(* Logix 5000 project; controller PLC_MCC1300_75F1 vendor 1 type 14 code 166 rev 32.11; software revision 32.04; part 16 of 83 *)
(* tags used below, declared in another part *)
   M302SpeedUp : MAC_SpeedUp;
   TMP_d : DINT;
   TMP_xPositioning : BOOL;
   TMP_xReverse : BOOL;
   TMP_xRun : BOOL;
   xAlwaysOFF : BOOL;
   Z300_Conveyor : UDT_StandConv[29];
   Z300_Conveyor_Conf : UDT_Conveyor_Config[29];
   Z300_Conveyor_HMW : MAC_Conveyor_ZC_HMW[29];
   Z300_Conveyor_IN_MOTION : MAC_Conveyor_ZC_IN_MOTION[29];
   Z301_HMR : MAC_Zone_ML_HMR;
(* CommandLogic, continued *)

ROUTINE M307AM2_Conveyor_Output   (* ladder *)
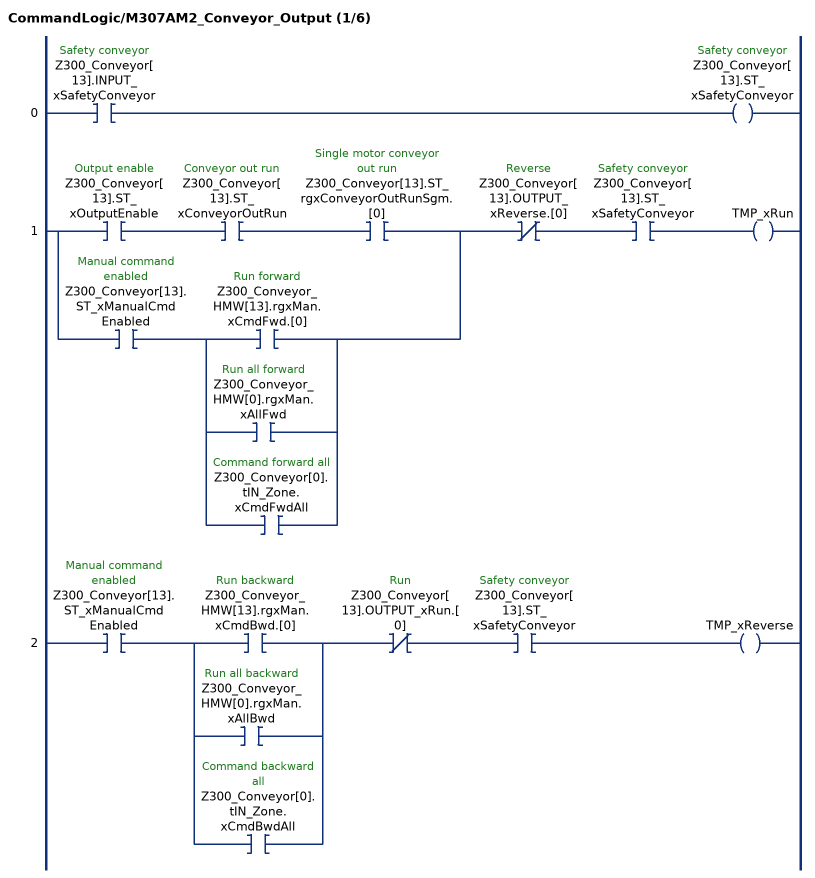
   0: XIC(Z300_Conveyor[13].INPUT_xSafetyConveyor)OTE(Z300_Conveyor[13].ST_xSafetyConveyor);
   1: [XIC(Z300_Conveyor[13].ST_xOutputEnable) XIC(Z300_Conveyor[13].ST_xConveyorOutRun) XIC(Z300_Conveyor[13].ST_rgxConveyorOutRunSgm.[0]) ,XIC(Z300_Conveyor[13].ST_xManualCmdEnabled) [XIC(Z300_Conveyor_HMW[13].rgxMan.xCmdFwd.[0]) ,XIC(Z300_Conveyor_HMW[0].rgxMan.xAllFwd) ,XIC(Z300_Conveyor[0].tIN_Zone.xCmdFwdAll) ] ]XIO(Z300_Conveyor[13].OUTPUT_xReverse.[0])XIC(Z300_Conveyor[13].ST_xSafetyConveyor)OTE(TMP_xRun);
   2: XIC(Z300_Conveyor[13].ST_xManualCmdEnabled)[XIC(Z300_Conveyor_HMW[13].rgxMan.xCmdBwd.[0]) ,XIC(Z300_Conveyor_HMW[0].rgxMan.xAllBwd) ,XIC(Z300_Conveyor[0].tIN_Zone.xCmdBwdAll) ]XIO(Z300_Conveyor[13].OUTPUT_xRun.[0])XIC(Z300_Conveyor[13].ST_xSafetyConveyor)OTE(TMP_xReverse);
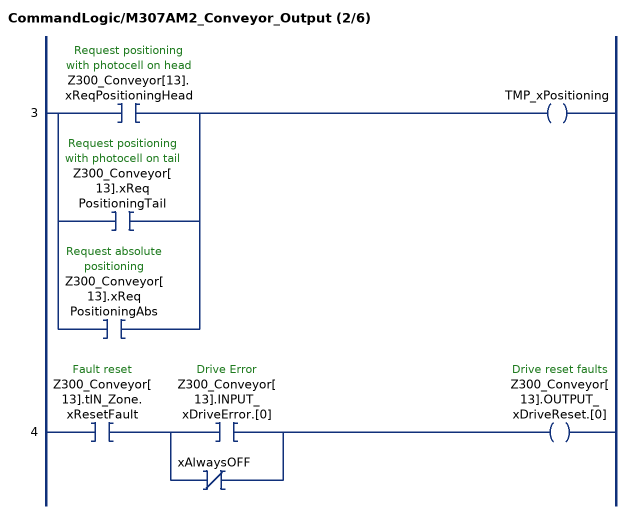
   3: [XIC(Z300_Conveyor[13].xReqPositioningHead) ,XIC(Z300_Conveyor[13].xReqPositioningTail) ,XIC(Z300_Conveyor[13].xReqPositioningAbs) ]OTE(TMP_xPositioning);
   4: XIC(Z300_Conveyor[13].tIN_Zone.xResetFault)[XIC(Z300_Conveyor[13].INPUT_xDriveError.[0]) ,XIO(xAlwaysOFF) ]OTE(Z300_Conveyor[13].OUTPUT_xDriveReset.[0]);
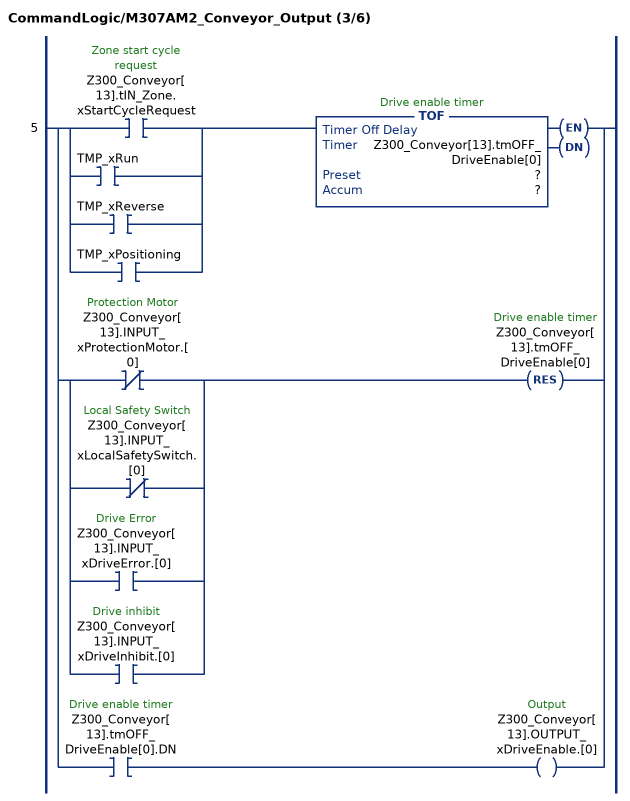
   5: [[XIC(Z300_Conveyor[13].tIN_Zone.xStartCycleRequest) ,XIC(TMP_xRun) ,XIC(TMP_xReverse) ,XIC(TMP_xPositioning) ] TOF(Z300_Conveyor[13].tmOFF_DriveEnable[0],?,?) ,[XIO(Z300_Conveyor[13].INPUT_xProtectionMotor.[0]) ,XIO(Z300_Conveyor[13].INPUT_xLocalSafetySwitch.[0]) ,XIC(Z300_Conveyor[13].INPUT_xDriveError.[0]) ,XIC(Z300_Conveyor[13].INPUT_xDriveInhibit.[0]) ] RES(Z300_Conveyor[13].tmOFF_DriveEnable[0]) ,XIC(Z300_Conveyor[13].tmOFF_DriveEnable[0].DN) OTE(Z300_Conveyor[13].OUTPUT_xDriveEnable.[0]) ];
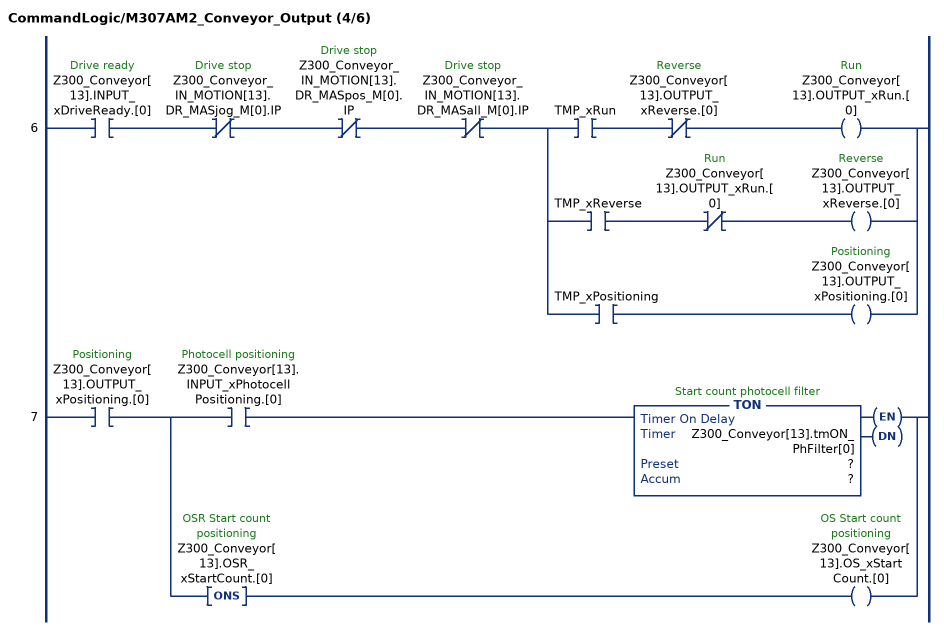
   6: XIC(Z300_Conveyor[13].INPUT_xDriveReady.[0])XIO(Z300_Conveyor_IN_MOTION[13].DR_MASjog_M[0].IP)XIO(Z300_Conveyor_IN_MOTION[13].DR_MASpos_M[0].IP)XIO(Z300_Conveyor_IN_MOTION[13].DR_MASall_M[0].IP)[XIC(TMP_xRun) XIO(Z300_Conveyor[13].OUTPUT_xReverse.[0]) OTE(Z300_Conveyor[13].OUTPUT_xRun.[0]) ,XIC(TMP_xReverse) XIO(Z300_Conveyor[13].OUTPUT_xRun.[0]) OTE(Z300_Conveyor[13].OUTPUT_xReverse.[0]) ,XIC(TMP_xPositioning) OTE(Z300_Conveyor[13].OUTPUT_xPositioning.[0]) ];
   7: XIC(Z300_Conveyor[13].OUTPUT_xPositioning.[0])[XIC(Z300_Conveyor[13].INPUT_xPhotocellPositioning.[0]) TON(Z300_Conveyor[13].tmON_PhFilter[0],?,?) ,ONS(Z300_Conveyor[13].OSR_xStartCount.[0]) OTE(Z300_Conveyor[13].OS_xStartCount.[0]) ];
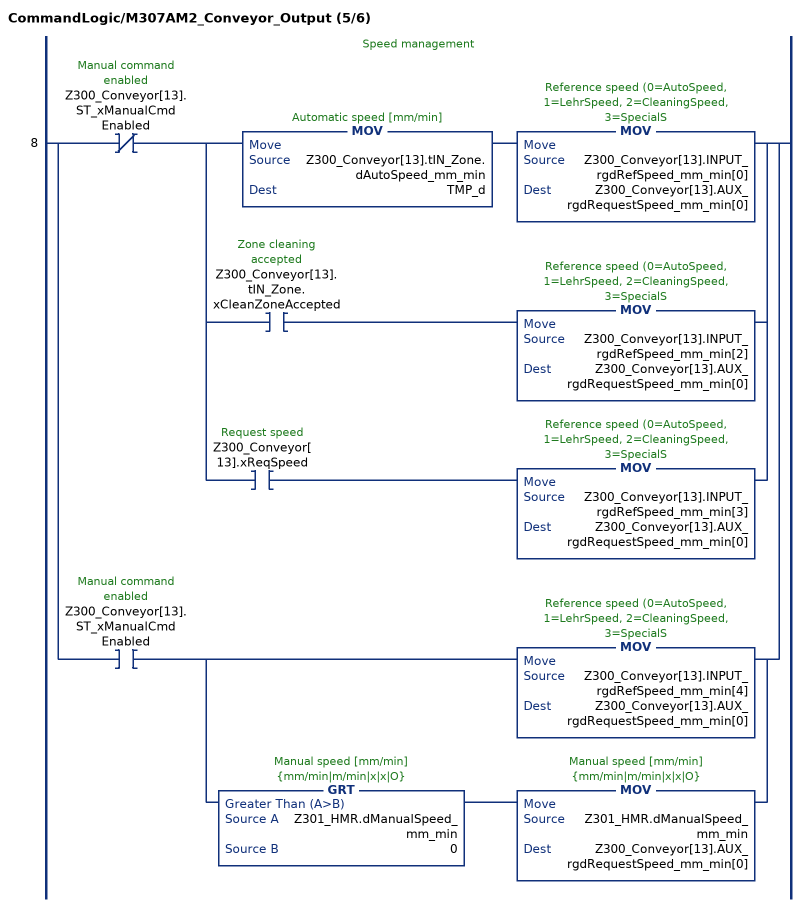
   // Speed management
   8: [XIO(Z300_Conveyor[13].ST_xManualCmdEnabled) [MOV(Z300_Conveyor[13].tIN_Zone.dAutoSpeed_mm_min,TMP_d) MOV(Z300_Conveyor[13].INPUT_rgdRefSpeed_mm_min[0],Z300_Conveyor[13].AUX_rgdRequestSpeed_mm_min[0]) ,XIC(Z300_Conveyor[13].tIN_Zone.xCleanZoneAccepted) MOV(Z300_Conveyor[13].INPUT_rgdRefSpeed_mm_min[2],Z300_Conveyor[13].AUX_rgdRequestSpeed_mm_min[0]) ,XIC(Z300_Conveyor[13].xReqSpeed) MOV(Z300_Conveyor[13].INPUT_rgdRefSpeed_mm_min[3],Z300_Conveyor[13].AUX_rgdRequestSpeed_mm_min[0]) ] ,XIC(Z300_Conveyor[13].ST_xManualCmdEnabled) [MOV(Z300_Conveyor[13].INPUT_rgdRefSpeed_mm_min[4],Z300_Conveyor[13].AUX_rgdRequestSpeed_mm_min[0]) ,GRT(Z301_HMR.dManualSpeed_mm_min,0) MOV(Z301_HMR.dManualSpeed_mm_min,Z300_Conveyor[13].AUX_rgdRequestSpeed_mm_min[0]) ] ];
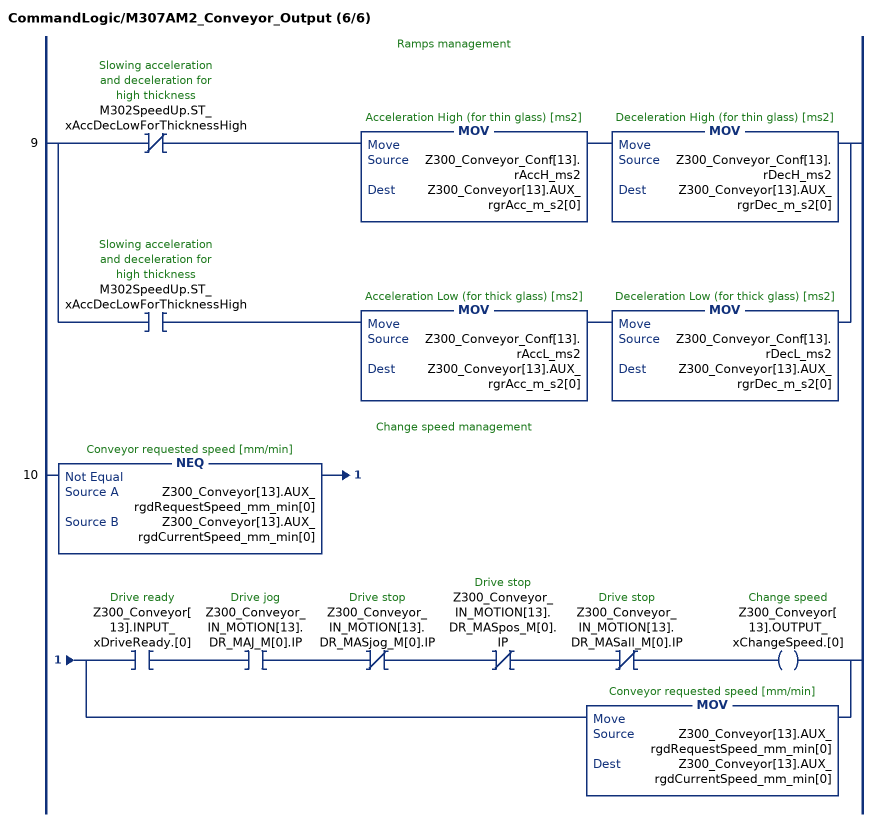
   // Ramps management
   9: [XIO(M302SpeedUp.ST_xAccDecLowForThicknessHigh) MOV(Z300_Conveyor_Conf[13].rAccH_ms2,Z300_Conveyor[13].AUX_rgrAcc_m_s2[0]) MOV(Z300_Conveyor_Conf[13].rDecH_ms2,Z300_Conveyor[13].AUX_rgrDec_m_s2[0]) ,XIC(M302SpeedUp.ST_xAccDecLowForThicknessHigh) MOV(Z300_Conveyor_Conf[13].rAccL_ms2,Z300_Conveyor[13].AUX_rgrAcc_m_s2[0]) MOV(Z300_Conveyor_Conf[13].rDecL_ms2,Z300_Conveyor[13].AUX_rgrDec_m_s2[0]) ];
   // Change speed management
   10: NEQ(Z300_Conveyor[13].AUX_rgdRequestSpeed_mm_min[0],Z300_Conveyor[13].AUX_rgdCurrentSpeed_mm_min[0])[XIC(Z300_Conveyor[13].INPUT_xDriveReady.[0]) XIC(Z300_Conveyor_IN_MOTION[13].DR_MAJ_M[0].IP) XIO(Z300_Conveyor_IN_MOTION[13].DR_MASjog_M[0].IP) XIO(Z300_Conveyor_IN_MOTION[13].DR_MASpos_M[0].IP) XIO(Z300_Conveyor_IN_MOTION[13].DR_MASall_M[0].IP) OTE(Z300_Conveyor[13].OUTPUT_xChangeSpeed.[0]) ,MOV(Z300_Conveyor[13].AUX_rgdRequestSpeed_mm_min[0],Z300_Conveyor[13].AUX_rgdCurrentSpeed_mm_min[0]) ];
END_ROUTINE

ROUTINE M307AM3_Conveyor_Output   (* ladder *)
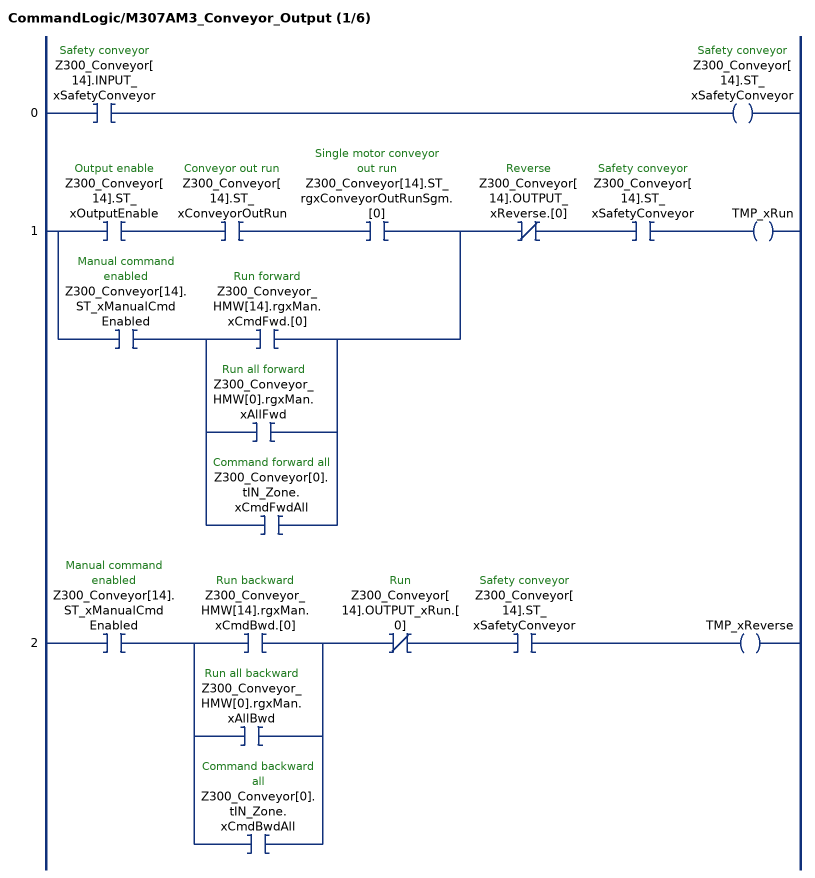
   0: XIC(Z300_Conveyor[14].INPUT_xSafetyConveyor)OTE(Z300_Conveyor[14].ST_xSafetyConveyor);
   1: [XIC(Z300_Conveyor[14].ST_xOutputEnable) XIC(Z300_Conveyor[14].ST_xConveyorOutRun) XIC(Z300_Conveyor[14].ST_rgxConveyorOutRunSgm.[0]) ,XIC(Z300_Conveyor[14].ST_xManualCmdEnabled) [XIC(Z300_Conveyor_HMW[14].rgxMan.xCmdFwd.[0]) ,XIC(Z300_Conveyor_HMW[0].rgxMan.xAllFwd) ,XIC(Z300_Conveyor[0].tIN_Zone.xCmdFwdAll) ] ]XIO(Z300_Conveyor[14].OUTPUT_xReverse.[0])XIC(Z300_Conveyor[14].ST_xSafetyConveyor)OTE(TMP_xRun);
   2: XIC(Z300_Conveyor[14].ST_xManualCmdEnabled)[XIC(Z300_Conveyor_HMW[14].rgxMan.xCmdBwd.[0]) ,XIC(Z300_Conveyor_HMW[0].rgxMan.xAllBwd) ,XIC(Z300_Conveyor[0].tIN_Zone.xCmdBwdAll) ]XIO(Z300_Conveyor[14].OUTPUT_xRun.[0])XIC(Z300_Conveyor[14].ST_xSafetyConveyor)OTE(TMP_xReverse);
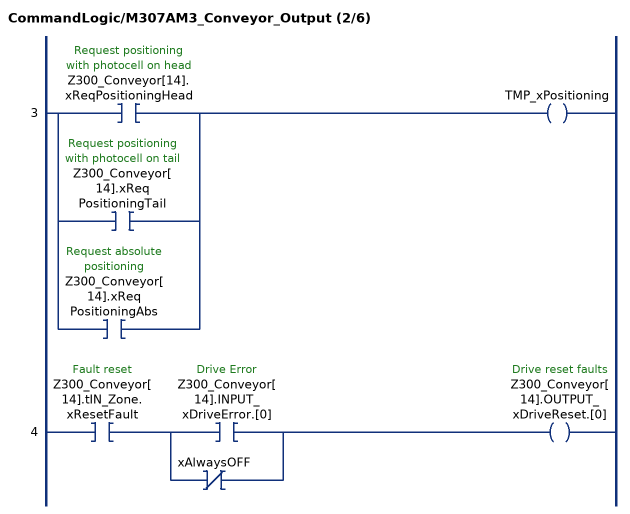
   3: [XIC(Z300_Conveyor[14].xReqPositioningHead) ,XIC(Z300_Conveyor[14].xReqPositioningTail) ,XIC(Z300_Conveyor[14].xReqPositioningAbs) ]OTE(TMP_xPositioning);
   4: XIC(Z300_Conveyor[14].tIN_Zone.xResetFault)[XIC(Z300_Conveyor[14].INPUT_xDriveError.[0]) ,XIO(xAlwaysOFF) ]OTE(Z300_Conveyor[14].OUTPUT_xDriveReset.[0]);
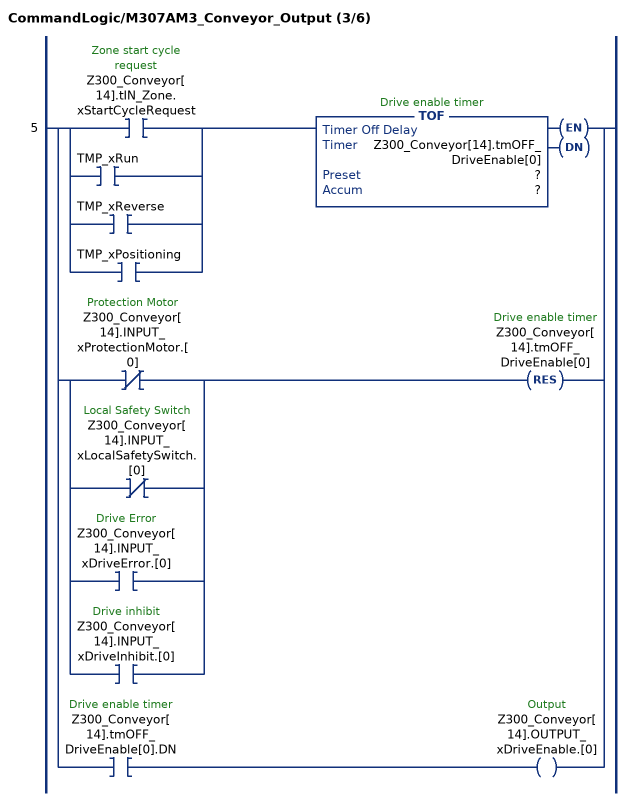
   5: [[XIC(Z300_Conveyor[14].tIN_Zone.xStartCycleRequest) ,XIC(TMP_xRun) ,XIC(TMP_xReverse) ,XIC(TMP_xPositioning) ] TOF(Z300_Conveyor[14].tmOFF_DriveEnable[0],?,?) ,[XIO(Z300_Conveyor[14].INPUT_xProtectionMotor.[0]) ,XIO(Z300_Conveyor[14].INPUT_xLocalSafetySwitch.[0]) ,XIC(Z300_Conveyor[14].INPUT_xDriveError.[0]) ,XIC(Z300_Conveyor[14].INPUT_xDriveInhibit.[0]) ] RES(Z300_Conveyor[14].tmOFF_DriveEnable[0]) ,XIC(Z300_Conveyor[14].tmOFF_DriveEnable[0].DN) OTE(Z300_Conveyor[14].OUTPUT_xDriveEnable.[0]) ];
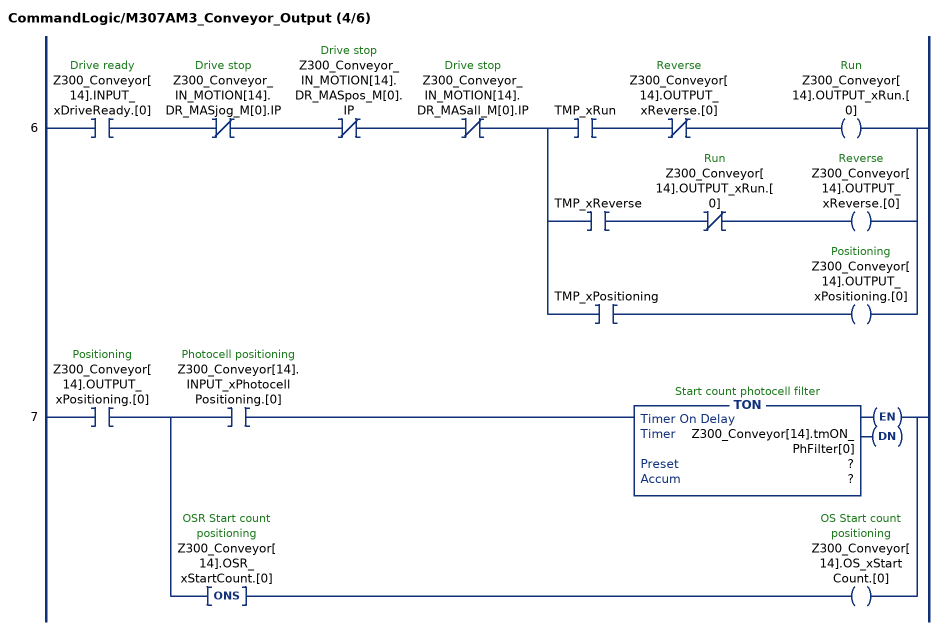
   6: XIC(Z300_Conveyor[14].INPUT_xDriveReady.[0])XIO(Z300_Conveyor_IN_MOTION[14].DR_MASjog_M[0].IP)XIO(Z300_Conveyor_IN_MOTION[14].DR_MASpos_M[0].IP)XIO(Z300_Conveyor_IN_MOTION[14].DR_MASall_M[0].IP)[XIC(TMP_xRun) XIO(Z300_Conveyor[14].OUTPUT_xReverse.[0]) OTE(Z300_Conveyor[14].OUTPUT_xRun.[0]) ,XIC(TMP_xReverse) XIO(Z300_Conveyor[14].OUTPUT_xRun.[0]) OTE(Z300_Conveyor[14].OUTPUT_xReverse.[0]) ,XIC(TMP_xPositioning) OTE(Z300_Conveyor[14].OUTPUT_xPositioning.[0]) ];
   7: XIC(Z300_Conveyor[14].OUTPUT_xPositioning.[0])[XIC(Z300_Conveyor[14].INPUT_xPhotocellPositioning.[0]) TON(Z300_Conveyor[14].tmON_PhFilter[0],?,?) ,ONS(Z300_Conveyor[14].OSR_xStartCount.[0]) OTE(Z300_Conveyor[14].OS_xStartCount.[0]) ];
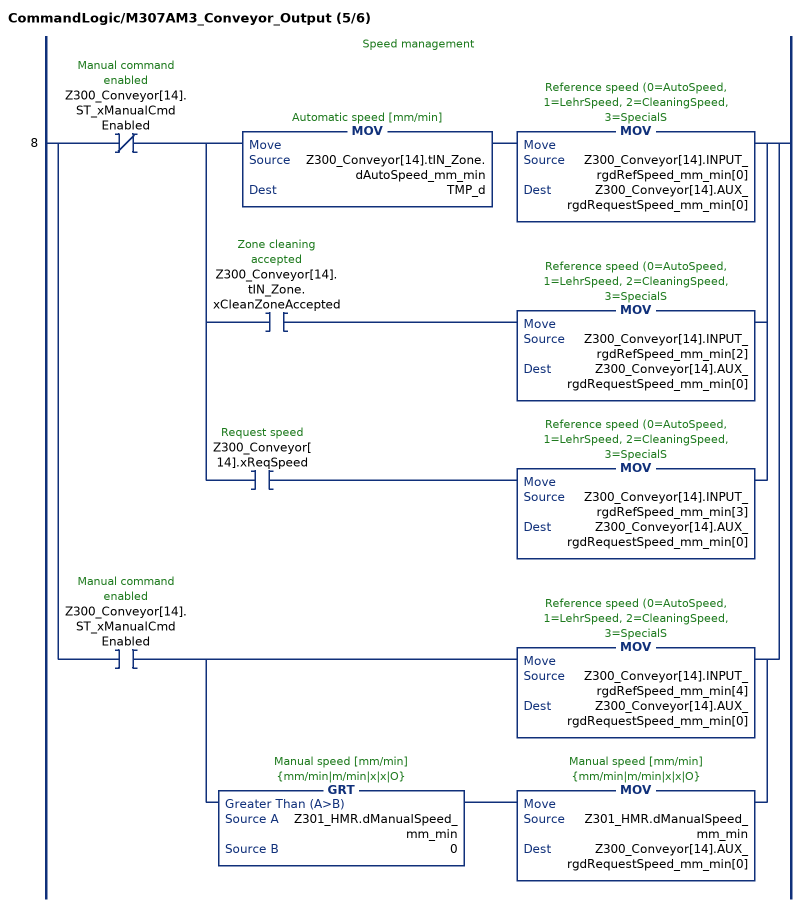
   // Speed management
   8: [XIO(Z300_Conveyor[14].ST_xManualCmdEnabled) [MOV(Z300_Conveyor[14].tIN_Zone.dAutoSpeed_mm_min,TMP_d) MOV(Z300_Conveyor[14].INPUT_rgdRefSpeed_mm_min[0],Z300_Conveyor[14].AUX_rgdRequestSpeed_mm_min[0]) ,XIC(Z300_Conveyor[14].tIN_Zone.xCleanZoneAccepted) MOV(Z300_Conveyor[14].INPUT_rgdRefSpeed_mm_min[2],Z300_Conveyor[14].AUX_rgdRequestSpeed_mm_min[0]) ,XIC(Z300_Conveyor[14].xReqSpeed) MOV(Z300_Conveyor[14].INPUT_rgdRefSpeed_mm_min[3],Z300_Conveyor[14].AUX_rgdRequestSpeed_mm_min[0]) ] ,XIC(Z300_Conveyor[14].ST_xManualCmdEnabled) [MOV(Z300_Conveyor[14].INPUT_rgdRefSpeed_mm_min[4],Z300_Conveyor[14].AUX_rgdRequestSpeed_mm_min[0]) ,GRT(Z301_HMR.dManualSpeed_mm_min,0) MOV(Z301_HMR.dManualSpeed_mm_min,Z300_Conveyor[14].AUX_rgdRequestSpeed_mm_min[0]) ] ];
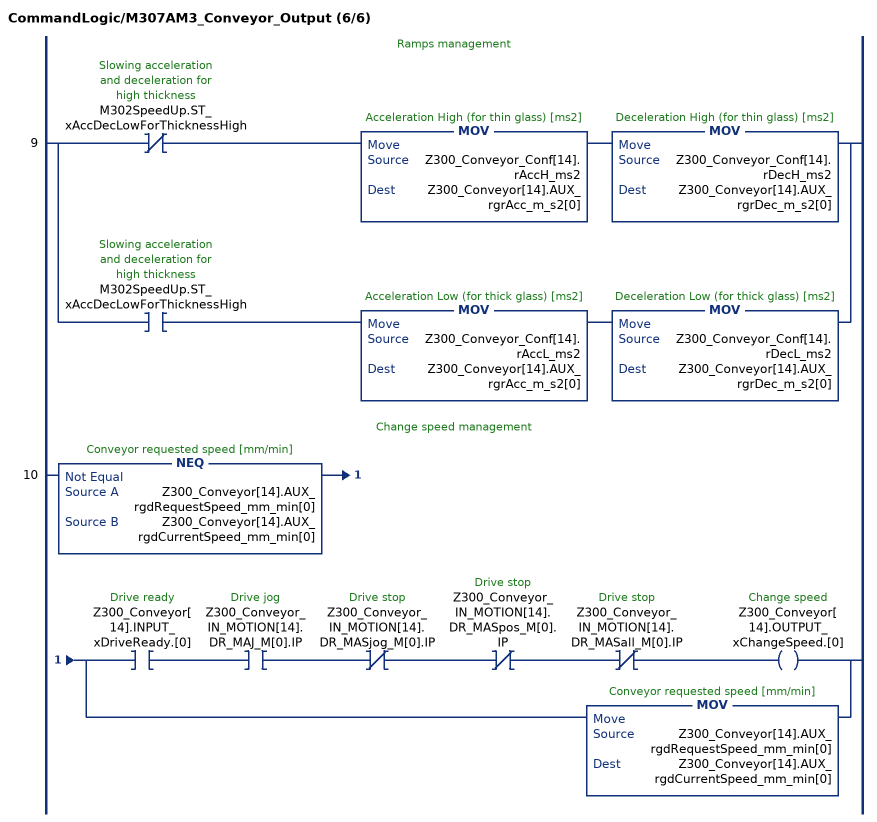
   // Ramps management
   9: [XIO(M302SpeedUp.ST_xAccDecLowForThicknessHigh) MOV(Z300_Conveyor_Conf[14].rAccH_ms2,Z300_Conveyor[14].AUX_rgrAcc_m_s2[0]) MOV(Z300_Conveyor_Conf[14].rDecH_ms2,Z300_Conveyor[14].AUX_rgrDec_m_s2[0]) ,XIC(M302SpeedUp.ST_xAccDecLowForThicknessHigh) MOV(Z300_Conveyor_Conf[14].rAccL_ms2,Z300_Conveyor[14].AUX_rgrAcc_m_s2[0]) MOV(Z300_Conveyor_Conf[14].rDecL_ms2,Z300_Conveyor[14].AUX_rgrDec_m_s2[0]) ];
   // Change speed management
   10: NEQ(Z300_Conveyor[14].AUX_rgdRequestSpeed_mm_min[0],Z300_Conveyor[14].AUX_rgdCurrentSpeed_mm_min[0])[XIC(Z300_Conveyor[14].INPUT_xDriveReady.[0]) XIC(Z300_Conveyor_IN_MOTION[14].DR_MAJ_M[0].IP) XIO(Z300_Conveyor_IN_MOTION[14].DR_MASjog_M[0].IP) XIO(Z300_Conveyor_IN_MOTION[14].DR_MASpos_M[0].IP) XIO(Z300_Conveyor_IN_MOTION[14].DR_MASall_M[0].IP) OTE(Z300_Conveyor[14].OUTPUT_xChangeSpeed.[0]) ,MOV(Z300_Conveyor[14].AUX_rgdRequestSpeed_mm_min[0],Z300_Conveyor[14].AUX_rgdCurrentSpeed_mm_min[0]) ];
END_ROUTINE

ROUTINE M307AM4_Conveyor_Output   (* ladder *)
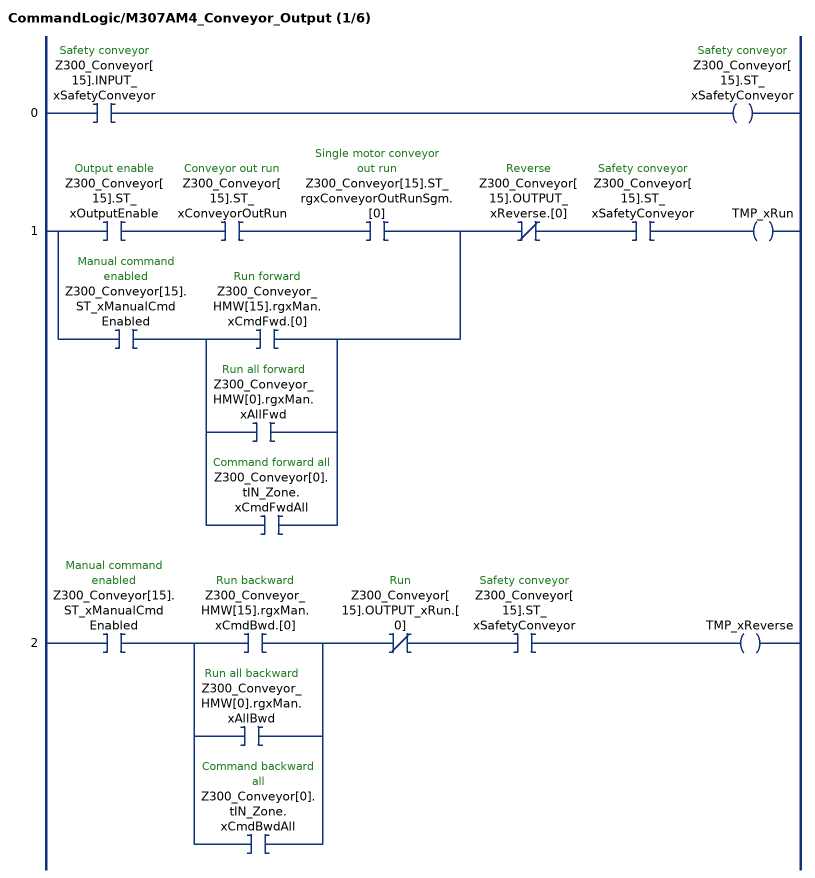
   0: XIC(Z300_Conveyor[15].INPUT_xSafetyConveyor)OTE(Z300_Conveyor[15].ST_xSafetyConveyor);
   1: [XIC(Z300_Conveyor[15].ST_xOutputEnable) XIC(Z300_Conveyor[15].ST_xConveyorOutRun) XIC(Z300_Conveyor[15].ST_rgxConveyorOutRunSgm.[0]) ,XIC(Z300_Conveyor[15].ST_xManualCmdEnabled) [XIC(Z300_Conveyor_HMW[15].rgxMan.xCmdFwd.[0]) ,XIC(Z300_Conveyor_HMW[0].rgxMan.xAllFwd) ,XIC(Z300_Conveyor[0].tIN_Zone.xCmdFwdAll) ] ]XIO(Z300_Conveyor[15].OUTPUT_xReverse.[0])XIC(Z300_Conveyor[15].ST_xSafetyConveyor)OTE(TMP_xRun);
   2: XIC(Z300_Conveyor[15].ST_xManualCmdEnabled)[XIC(Z300_Conveyor_HMW[15].rgxMan.xCmdBwd.[0]) ,XIC(Z300_Conveyor_HMW[0].rgxMan.xAllBwd) ,XIC(Z300_Conveyor[0].tIN_Zone.xCmdBwdAll) ]XIO(Z300_Conveyor[15].OUTPUT_xRun.[0])XIC(Z300_Conveyor[15].ST_xSafetyConveyor)OTE(TMP_xReverse);
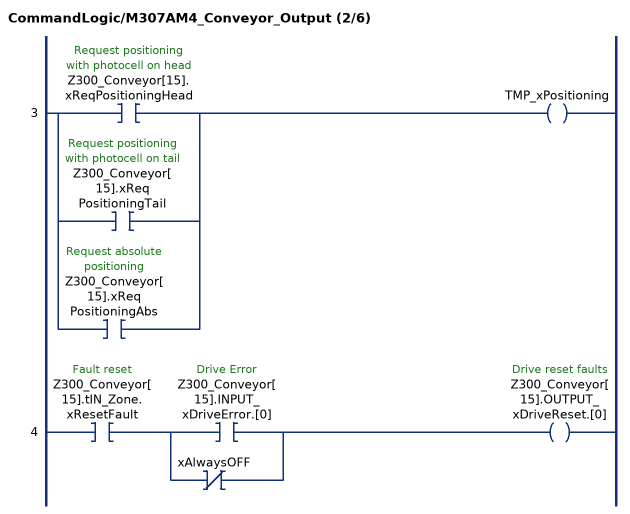
   3: [XIC(Z300_Conveyor[15].xReqPositioningHead) ,XIC(Z300_Conveyor[15].xReqPositioningTail) ,XIC(Z300_Conveyor[15].xReqPositioningAbs) ]OTE(TMP_xPositioning);
   4: XIC(Z300_Conveyor[15].tIN_Zone.xResetFault)[XIC(Z300_Conveyor[15].INPUT_xDriveError.[0]) ,XIO(xAlwaysOFF) ]OTE(Z300_Conveyor[15].OUTPUT_xDriveReset.[0]);
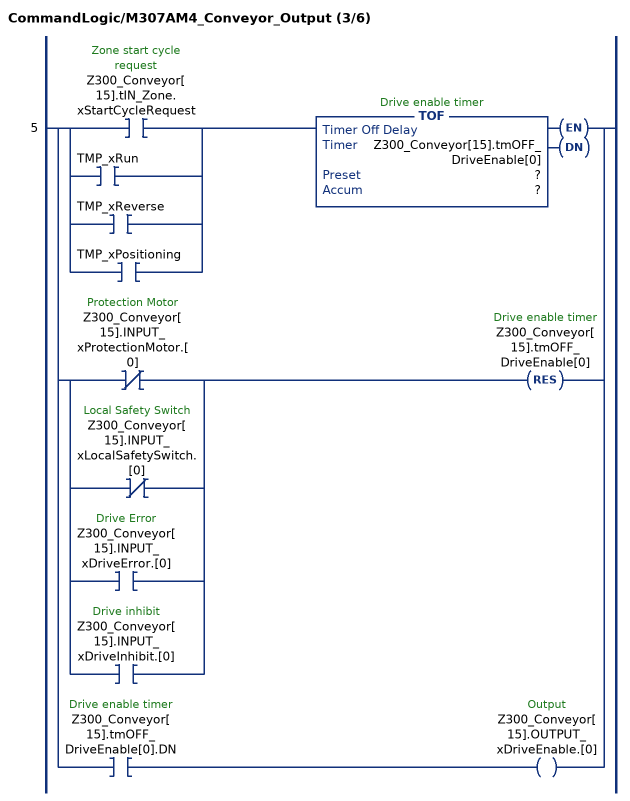
   5: [[XIC(Z300_Conveyor[15].tIN_Zone.xStartCycleRequest) ,XIC(TMP_xRun) ,XIC(TMP_xReverse) ,XIC(TMP_xPositioning) ] TOF(Z300_Conveyor[15].tmOFF_DriveEnable[0],?,?) ,[XIO(Z300_Conveyor[15].INPUT_xProtectionMotor.[0]) ,XIO(Z300_Conveyor[15].INPUT_xLocalSafetySwitch.[0]) ,XIC(Z300_Conveyor[15].INPUT_xDriveError.[0]) ,XIC(Z300_Conveyor[15].INPUT_xDriveInhibit.[0]) ] RES(Z300_Conveyor[15].tmOFF_DriveEnable[0]) ,XIC(Z300_Conveyor[15].tmOFF_DriveEnable[0].DN) OTE(Z300_Conveyor[15].OUTPUT_xDriveEnable.[0]) ];
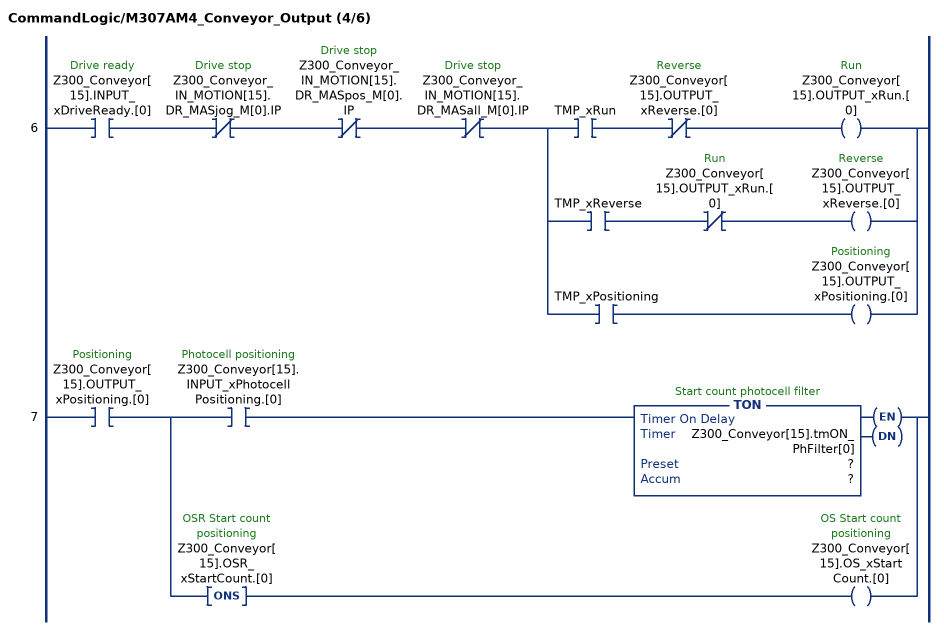
   6: XIC(Z300_Conveyor[15].INPUT_xDriveReady.[0])XIO(Z300_Conveyor_IN_MOTION[15].DR_MASjog_M[0].IP)XIO(Z300_Conveyor_IN_MOTION[15].DR_MASpos_M[0].IP)XIO(Z300_Conveyor_IN_MOTION[15].DR_MASall_M[0].IP)[XIC(TMP_xRun) XIO(Z300_Conveyor[15].OUTPUT_xReverse.[0]) OTE(Z300_Conveyor[15].OUTPUT_xRun.[0]) ,XIC(TMP_xReverse) XIO(Z300_Conveyor[15].OUTPUT_xRun.[0]) OTE(Z300_Conveyor[15].OUTPUT_xReverse.[0]) ,XIC(TMP_xPositioning) OTE(Z300_Conveyor[15].OUTPUT_xPositioning.[0]) ];
   7: XIC(Z300_Conveyor[15].OUTPUT_xPositioning.[0])[XIC(Z300_Conveyor[15].INPUT_xPhotocellPositioning.[0]) TON(Z300_Conveyor[15].tmON_PhFilter[0],?,?) ,ONS(Z300_Conveyor[15].OSR_xStartCount.[0]) OTE(Z300_Conveyor[15].OS_xStartCount.[0]) ];
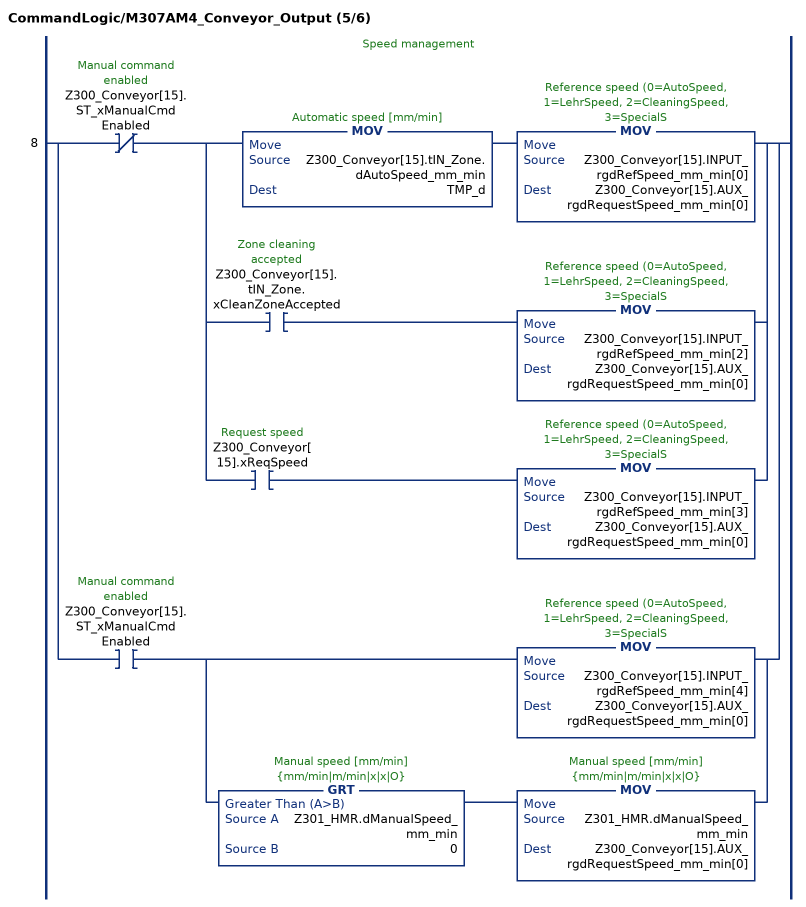
   // Speed management
   8: [XIO(Z300_Conveyor[15].ST_xManualCmdEnabled) [MOV(Z300_Conveyor[15].tIN_Zone.dAutoSpeed_mm_min,TMP_d) MOV(Z300_Conveyor[15].INPUT_rgdRefSpeed_mm_min[0],Z300_Conveyor[15].AUX_rgdRequestSpeed_mm_min[0]) ,XIC(Z300_Conveyor[15].tIN_Zone.xCleanZoneAccepted) MOV(Z300_Conveyor[15].INPUT_rgdRefSpeed_mm_min[2],Z300_Conveyor[15].AUX_rgdRequestSpeed_mm_min[0]) ,XIC(Z300_Conveyor[15].xReqSpeed) MOV(Z300_Conveyor[15].INPUT_rgdRefSpeed_mm_min[3],Z300_Conveyor[15].AUX_rgdRequestSpeed_mm_min[0]) ] ,XIC(Z300_Conveyor[15].ST_xManualCmdEnabled) [MOV(Z300_Conveyor[15].INPUT_rgdRefSpeed_mm_min[4],Z300_Conveyor[15].AUX_rgdRequestSpeed_mm_min[0]) ,GRT(Z301_HMR.dManualSpeed_mm_min,0) MOV(Z301_HMR.dManualSpeed_mm_min,Z300_Conveyor[15].AUX_rgdRequestSpeed_mm_min[0]) ] ];
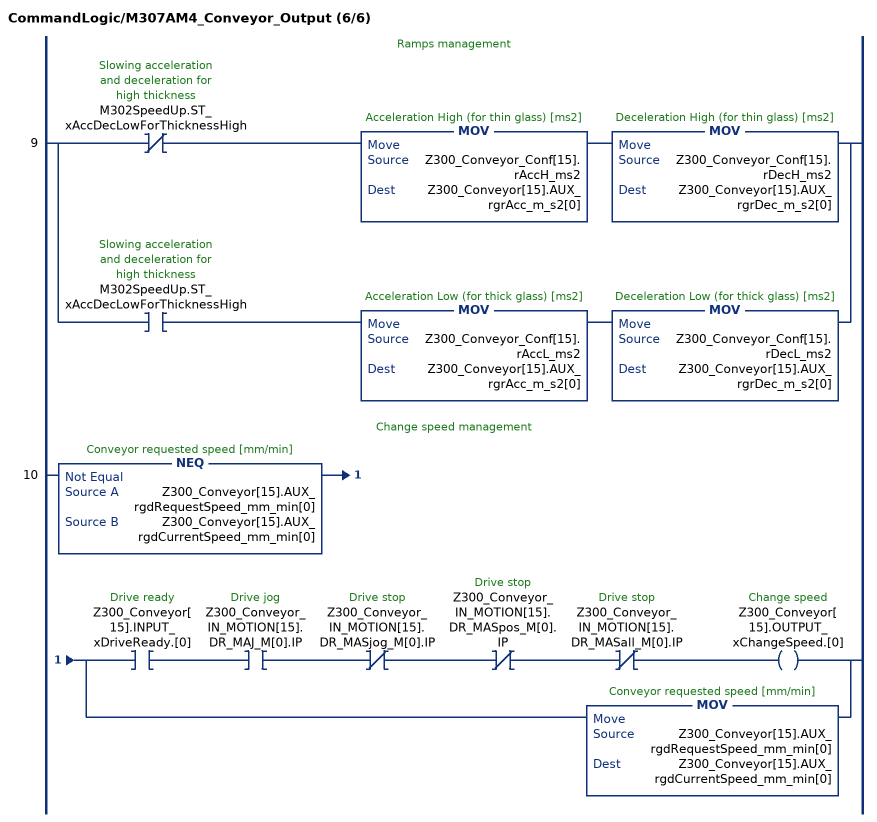
   // Ramps management
   9: [XIO(M302SpeedUp.ST_xAccDecLowForThicknessHigh) MOV(Z300_Conveyor_Conf[15].rAccH_ms2,Z300_Conveyor[15].AUX_rgrAcc_m_s2[0]) MOV(Z300_Conveyor_Conf[15].rDecH_ms2,Z300_Conveyor[15].AUX_rgrDec_m_s2[0]) ,XIC(M302SpeedUp.ST_xAccDecLowForThicknessHigh) MOV(Z300_Conveyor_Conf[15].rAccL_ms2,Z300_Conveyor[15].AUX_rgrAcc_m_s2[0]) MOV(Z300_Conveyor_Conf[15].rDecL_ms2,Z300_Conveyor[15].AUX_rgrDec_m_s2[0]) ];
   // Change speed management
   10: NEQ(Z300_Conveyor[15].AUX_rgdRequestSpeed_mm_min[0],Z300_Conveyor[15].AUX_rgdCurrentSpeed_mm_min[0])[XIC(Z300_Conveyor[15].INPUT_xDriveReady.[0]) XIC(Z300_Conveyor_IN_MOTION[15].DR_MAJ_M[0].IP) XIO(Z300_Conveyor_IN_MOTION[15].DR_MASjog_M[0].IP) XIO(Z300_Conveyor_IN_MOTION[15].DR_MASpos_M[0].IP) XIO(Z300_Conveyor_IN_MOTION[15].DR_MASall_M[0].IP) OTE(Z300_Conveyor[15].OUTPUT_xChangeSpeed.[0]) ,MOV(Z300_Conveyor[15].AUX_rgdRequestSpeed_mm_min[0],Z300_Conveyor[15].AUX_rgdCurrentSpeed_mm_min[0]) ];
END_ROUTINE
